(* Logix 5000 project; controller FV vendor 1 type 14 code 217 rev 31.11; software revision 31.00; part 37 of 63 *)
(* tags used below, declared in another part *)
   CWD : CHECKWORD_FLAGS;
   Dummy : BOOL;
   FV_bit_to_clear : DINT;
   FV_data_file_address : INT;
   FV_FV10C : PlantItem;   // FV10C
   FV_FV10J : PlantItem;   // FV10J
   FV_FV11C : PlantItem;   // FV11C
   FV_FV11J : PlantItem;   // FV11J
   FV_FV12C : PlantItem;   // FV12C
   FV_FV12J : PlantItem;   // FV12J
   FV_FV13C : PlantItem;   // FV13C
   FV_FV13J : PlantItem;   // FV13J
   FV_FV14C : PlantItem;   // FV14C
   FV_FV14J : PlantItem;   // FV14J
   FV_FV15C : PlantItem;   // FV15C
   FV_FV15J : PlantItem;   // FV15J
   FV_FV16C : PlantItem;   // FV16C
   FV_FV16J : PlantItem;   // FV16J
   FV_FV17C : PlantItem;   // FV17C
   FV_FV17J : PlantItem;   // FV17J
   FV_FV18C : PlantItem;   // FV18C
   FV_FV18J : PlantItem;   // FV18J
   FV_FV19C : PlantItem;   // FV19C
   FV_FV19J : PlantItem;   // FV19J
   FV_FV1C : PlantItem;   // FV1C
   FV_FV1J : PlantItem;   // FV1J
   FV_FV20C : PlantItem;   // FV20C
   FV_FV20J : PlantItem;   // FV20J
   FV_FV21C : PlantItem;   // FV21C
   FV_FV21J : PlantItem;   // FV21J
   FV_FV22C : PlantItem;   // FV22C
   FV_FV22J : PlantItem;   // FV22J
   FV_FV23C : PlantItem;   // FV23C
   FV_FV23J : PlantItem;   // FV23J
   FV_FV24C : PlantItem;   // FV24C
   FV_FV24J : PlantItem;   // FV24J
   FV_FV25C : PlantItem;   // FV25C
   FV_FV25J : PlantItem;   // FV25J
   FV_FV26C : PlantItem;   // FV26C
   FV_FV26J : PlantItem;   // FV26J
   FV_FV27C : PlantItem;   // FV27C
   FV_FV27J : PlantItem;   // FV27J
   FV_FV28C : PlantItem;   // FV28C
   FV_FV28J : PlantItem;   // FV28J
   FV_FV29C : PlantItem;   // FV29C
   FV_FV29J : PlantItem;   // FV29J
   FV_FV2C : PlantItem;   // FV2C
   FV_FV2J : PlantItem;   // FV2J
   FV_FV30C : PlantItem;   // FV30C
   FV_FV30J : PlantItem;   // FV30J
   FV_FV31C : PlantItem;   // FV31C
   FV_FV31J : PlantItem;   // FV31J
   FV_FV3C : PlantItem;   // FV3C
   FV_FV3J : PlantItem;   // FV3J
   FV_FV4C : PlantItem;   // FV4C
   FV_FV4J : PlantItem;   // FV4J
   FV_FV5C : PlantItem;   // FV5C
   FV_FV5J : PlantItem;   // FV5J
   FV_FV6C : PlantItem;   // FV6C
   FV_FV6J : PlantItem;   // FV6J
   FV_FV7C : PlantItem;   // FV7C
   FV_FV7J : PlantItem;   // FV7J
   FV_FV8C : PlantItem;   // FV8C
   FV_FV8J : PlantItem;   // FV8J
   FV_FV9C : PlantItem;   // FV9C
   FV_FV9J : PlantItem;   // FV9J
   FV_N110 : INT[255];   // FV DATA 0 CURRENT FV DATA
   FV_N111 : INT[50];   // FV1, CURRENT FV DATA
   FV_N112 : INT[50];   // FV2, CURRENT FV DATA
   FV_N113 : INT[50];   // FV3, CURRENT FV DATA
   FV_N114 : INT[50];   // FV4, CURRENT FV DATA
   FV_N115 : INT[50];   // FV5, CURRENT FV DATA
   FV_N116 : INT[50];   // FV6, CURRENT FV DATA
   FV_N117 : INT[50];   // FV7, CURRENT FV DATA
   FV_N118 : INT[50];   // FV8, CURRENT FV DATA
   FV_N119 : INT[50];   // FV9, CURRENT FV DATA
   FV_N120 : INT[50];   // FV10, CURRENT FV DATA
   FV_N121 : INT[50];   // FV11, CURRENT FV DATA
   FV_N122 : INT[50];   // FV12, CURRENT FV DATA
   FV_N123 : INT[50];   // FV13, CURRENT FV DATA
   FV_N124 : INT[50];   // FV14, CURRENT FV DATA
   FV_N125 : INT[50];   // FV15, CURRENT FV DATA
   FV_N126 : INT[50];   // FV16, CURRENT FV DATA
   FV_N127 : INT[50];   // FV17, CURRENT FV DATA
   FV_N128 : INT[50];   // FV18, CURRENT FV DATA
   FV_N129 : INT[50];   // FV19, CURRENT FV DATA
   FV_N13 : INT[255];   // PLC>ME Inter PLC comms traf fic inbound
   FV_N130 : INT[50];   // FV20, CURRENT FV DATA
   FV_N131 : INT[50];   // FV21, CURRENT FV DATA
   FV_N132 : INT[50];   // FV22, CURRENT FV DATA
   FV_N133 : INT[50];   // FV23, CURRENT FV DATA
   FV_N134 : INT[50];   // FV24, CURRENT FV DATA
   FV_N135 : INT[50];   // FV25, CURRENT FV DATA
   FV_N136 : INT[50];   // YSV1, CURRENT FV DATA
   FV_N137 : INT[50];   // YSV2, CURRENT FV DATA
   FV_N138 : INT[50];   // YSV3, CURRENT FV DATA
   FV_N139 : INT[255];   // YST1
   FV_N140 : INT[255];   // YST2
   FV_N141 : INT[255];   // YSV1 DATA
   FV_N142 : INT[255];   // YSV2 DATA
   FV_N143 : INT[255];   // YSV3 DATA
   FV_N144 : INT[255];   // YST1 DATA
   FV_N145 : INT[255];   // YST2 DATA
   FV_N146 : INT[50];   // FV26, CURRENT FV DATA
   FV_N147 : INT[50];   // FV27, CURRENT FV DATA
   FV_N148 : INT[50];   // FV28, CURRENT FV DATA
   FV_N149 : INT[50];   // FV29, CURRENT FV DATA
   FV_N150 : INT[50];   // FV30, CURRENT FV DATA
   FV_N151 : INT[50];   // FV31, CURRENT FV DATA
   FV_N210 : INT[255];   // GLYCL_PTRS
   FV_word_offset : INT;
   FV_YSV1CV : PlantItem;   // YSV1CV
   FV_YSV1J : PlantItem;   // YSV1J
   FV_YSV2CV : PlantItem;   // YSV2CV
   FV_YSV2J : PlantItem;   // YSV2J
   FV_YSV3J : PlantItem;   // YSV3J
(* FV_Common, continued *)

ROUTINE FV_Clear_Flag_In_FV_Datafile   (* ladder *)
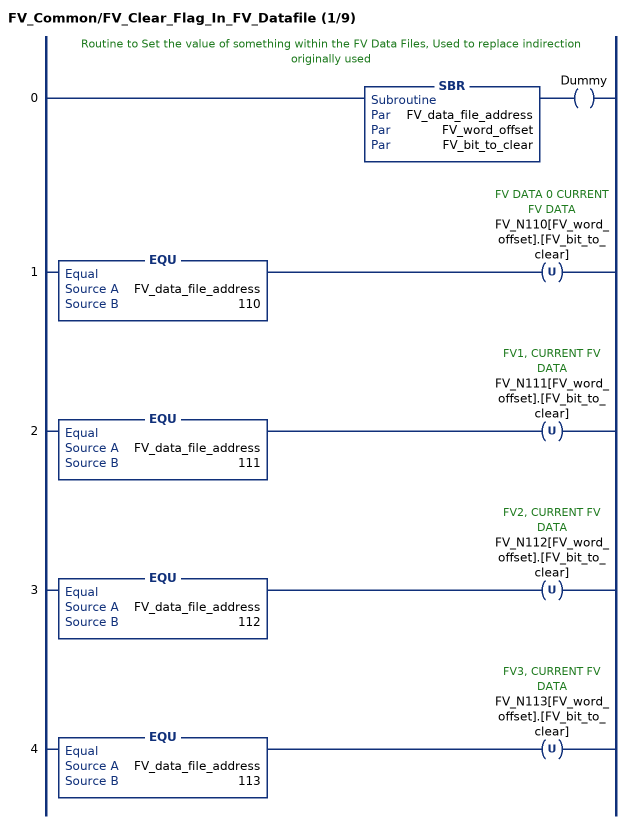
   // Routine to Set the value of something within the FV Data Files, Used to replace indirection originally used
   0: SBR(FV_data_file_address,FV_word_offset,FV_bit_to_clear)OTE(Dummy);
   1: EQU(FV_data_file_address,110)OTU(FV_N110[FV_word_offset].[FV_bit_to_clear]);
   2: EQU(FV_data_file_address,111)OTU(FV_N111[FV_word_offset].[FV_bit_to_clear]);
   3: EQU(FV_data_file_address,112)OTU(FV_N112[FV_word_offset].[FV_bit_to_clear]);
   4: EQU(FV_data_file_address,113)OTU(FV_N113[FV_word_offset].[FV_bit_to_clear]);
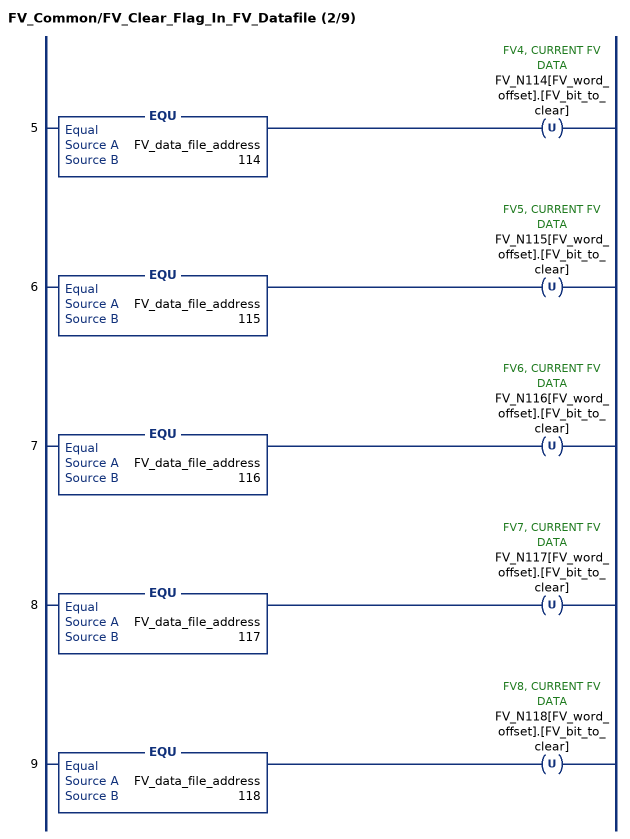
   5: EQU(FV_data_file_address,114)OTU(FV_N114[FV_word_offset].[FV_bit_to_clear]);
   6: EQU(FV_data_file_address,115)OTU(FV_N115[FV_word_offset].[FV_bit_to_clear]);
   7: EQU(FV_data_file_address,116)OTU(FV_N116[FV_word_offset].[FV_bit_to_clear]);
   8: EQU(FV_data_file_address,117)OTU(FV_N117[FV_word_offset].[FV_bit_to_clear]);
   9: EQU(FV_data_file_address,118)OTU(FV_N118[FV_word_offset].[FV_bit_to_clear]);
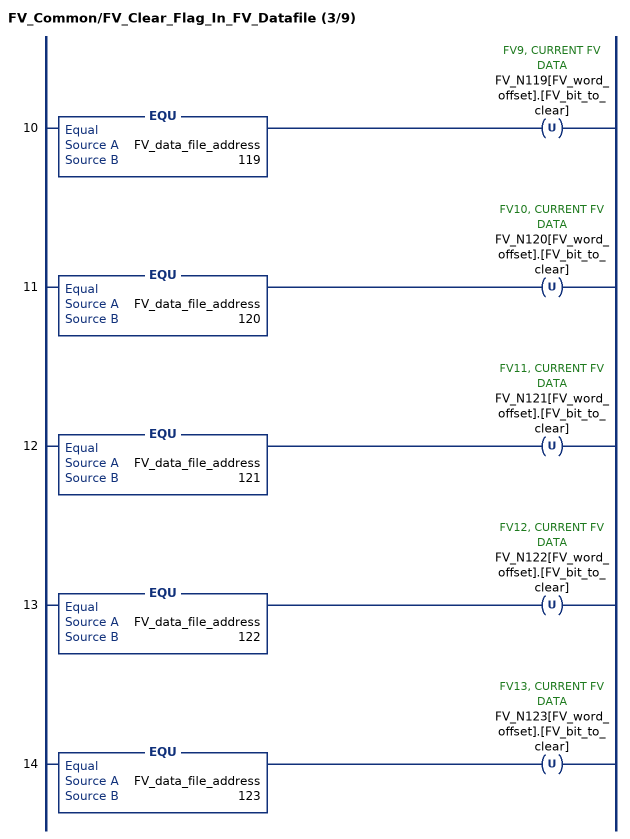
   10: EQU(FV_data_file_address,119)OTU(FV_N119[FV_word_offset].[FV_bit_to_clear]);
   11: EQU(FV_data_file_address,120)OTU(FV_N120[FV_word_offset].[FV_bit_to_clear]);
   12: EQU(FV_data_file_address,121)OTU(FV_N121[FV_word_offset].[FV_bit_to_clear]);
   13: EQU(FV_data_file_address,122)OTU(FV_N122[FV_word_offset].[FV_bit_to_clear]);
   14: EQU(FV_data_file_address,123)OTU(FV_N123[FV_word_offset].[FV_bit_to_clear]);
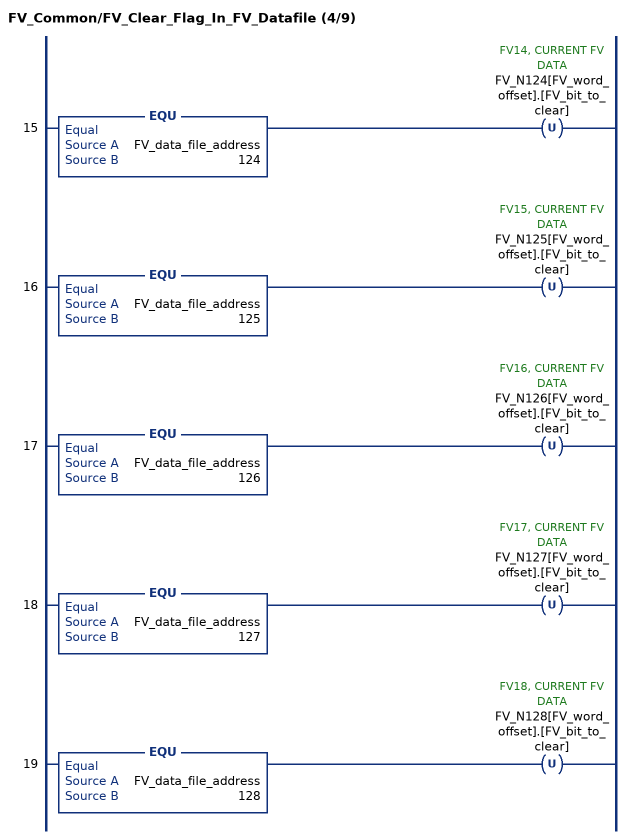
   15: EQU(FV_data_file_address,124)OTU(FV_N124[FV_word_offset].[FV_bit_to_clear]);
   16: EQU(FV_data_file_address,125)OTU(FV_N125[FV_word_offset].[FV_bit_to_clear]);
   17: EQU(FV_data_file_address,126)OTU(FV_N126[FV_word_offset].[FV_bit_to_clear]);
   18: EQU(FV_data_file_address,127)OTU(FV_N127[FV_word_offset].[FV_bit_to_clear]);
   19: EQU(FV_data_file_address,128)OTU(FV_N128[FV_word_offset].[FV_bit_to_clear]);
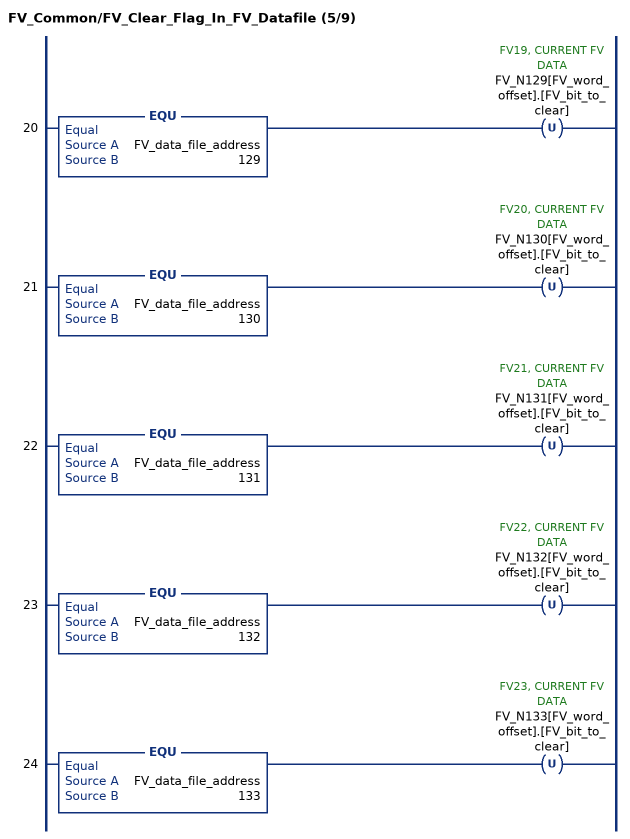
   20: EQU(FV_data_file_address,129)OTU(FV_N129[FV_word_offset].[FV_bit_to_clear]);
   21: EQU(FV_data_file_address,130)OTU(FV_N130[FV_word_offset].[FV_bit_to_clear]);
   22: EQU(FV_data_file_address,131)OTU(FV_N131[FV_word_offset].[FV_bit_to_clear]);
   23: EQU(FV_data_file_address,132)OTU(FV_N132[FV_word_offset].[FV_bit_to_clear]);
   24: EQU(FV_data_file_address,133)OTU(FV_N133[FV_word_offset].[FV_bit_to_clear]);
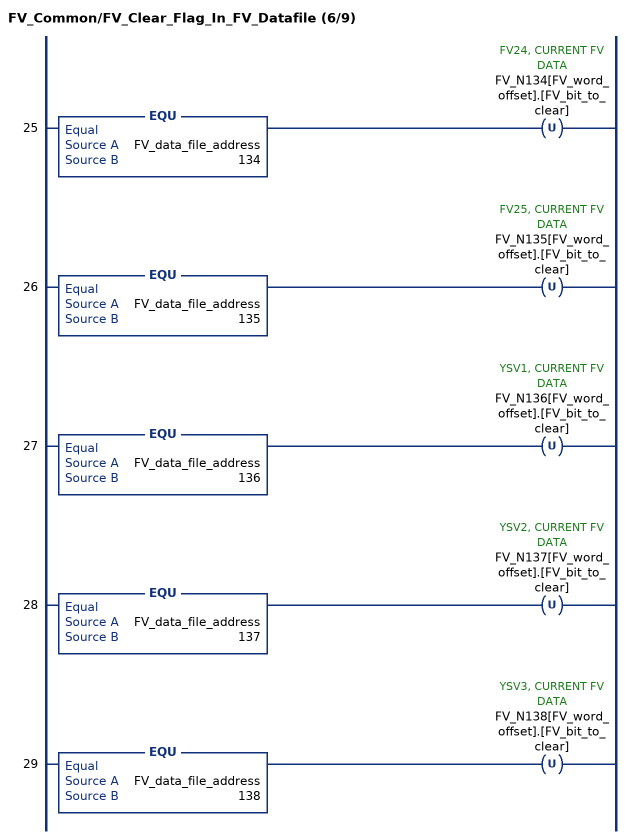
   25: EQU(FV_data_file_address,134)OTU(FV_N134[FV_word_offset].[FV_bit_to_clear]);
   26: EQU(FV_data_file_address,135)OTU(FV_N135[FV_word_offset].[FV_bit_to_clear]);
   27: EQU(FV_data_file_address,136)OTU(FV_N136[FV_word_offset].[FV_bit_to_clear]);
   28: EQU(FV_data_file_address,137)OTU(FV_N137[FV_word_offset].[FV_bit_to_clear]);
   29: EQU(FV_data_file_address,138)OTU(FV_N138[FV_word_offset].[FV_bit_to_clear]);
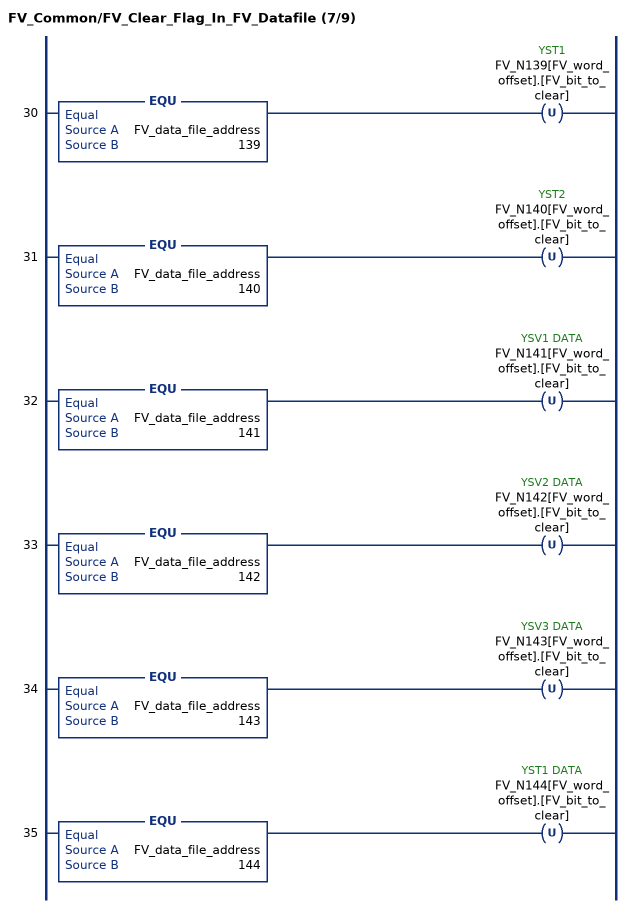
   30: EQU(FV_data_file_address,139)OTU(FV_N139[FV_word_offset].[FV_bit_to_clear]);
   31: EQU(FV_data_file_address,140)OTU(FV_N140[FV_word_offset].[FV_bit_to_clear]);
   32: EQU(FV_data_file_address,141)OTU(FV_N141[FV_word_offset].[FV_bit_to_clear]);
   33: EQU(FV_data_file_address,142)OTU(FV_N142[FV_word_offset].[FV_bit_to_clear]);
   34: EQU(FV_data_file_address,143)OTU(FV_N143[FV_word_offset].[FV_bit_to_clear]);
   35: EQU(FV_data_file_address,144)OTU(FV_N144[FV_word_offset].[FV_bit_to_clear]);
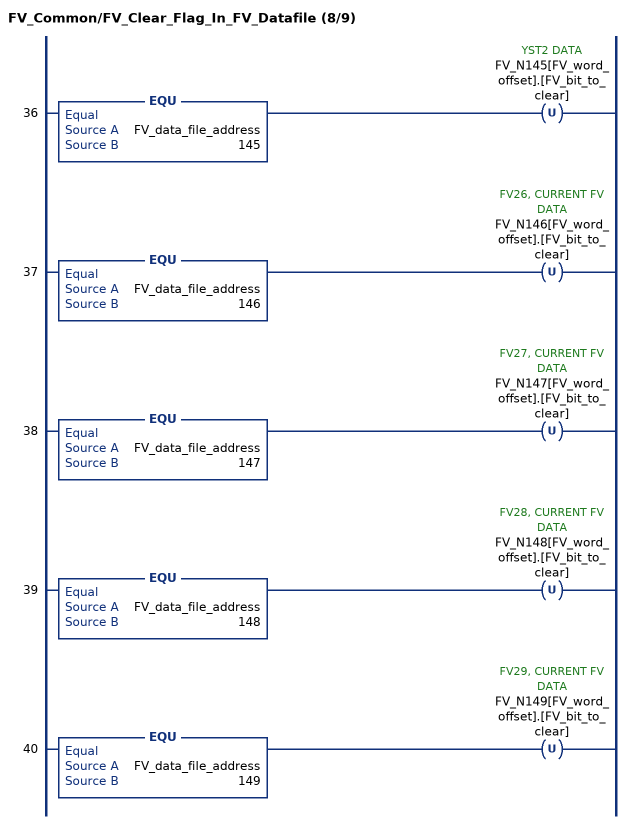
   36: EQU(FV_data_file_address,145)OTU(FV_N145[FV_word_offset].[FV_bit_to_clear]);
   37: EQU(FV_data_file_address,146)OTU(FV_N146[FV_word_offset].[FV_bit_to_clear]);
   38: EQU(FV_data_file_address,147)OTU(FV_N147[FV_word_offset].[FV_bit_to_clear]);
   39: EQU(FV_data_file_address,148)OTU(FV_N148[FV_word_offset].[FV_bit_to_clear]);
   40: EQU(FV_data_file_address,149)OTU(FV_N149[FV_word_offset].[FV_bit_to_clear]);
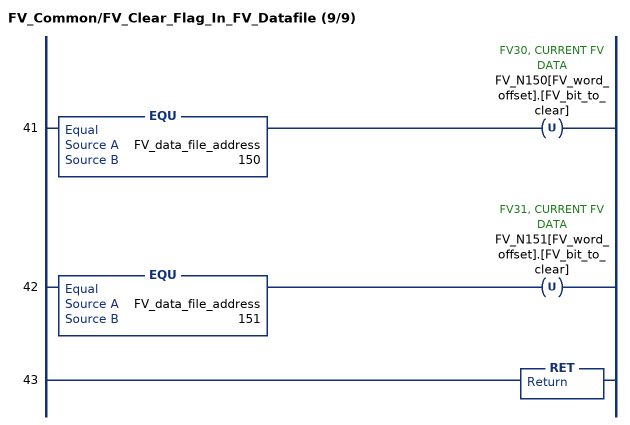
   41: EQU(FV_data_file_address,150)OTU(FV_N150[FV_word_offset].[FV_bit_to_clear]);
   42: EQU(FV_data_file_address,151)OTU(FV_N151[FV_word_offset].[FV_bit_to_clear]);
   43: RET();
END_ROUTINE

ROUTINE FV_COOLVLVOPN_111   (* ladder *)
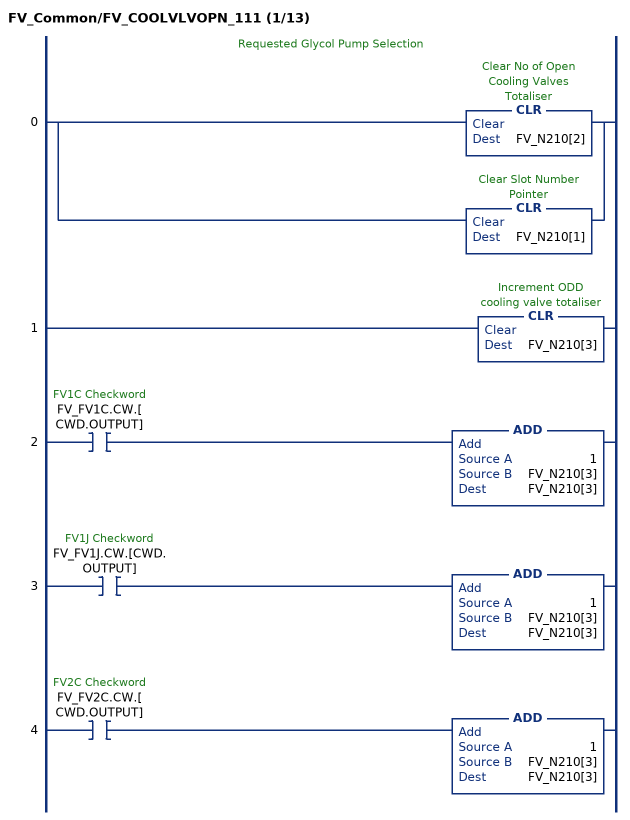
   // Requested Glycol Pump Selection
   0: [CLR(FV_N210[2]) ,CLR(FV_N210[1]) ];
   1: CLR(FV_N210[3]);
   2: XIC(FV_FV1C.CW.[CWD.OUTPUT])ADD(1,FV_N210[3],FV_N210[3]);
   3: XIC(FV_FV1J.CW.[CWD.OUTPUT])ADD(1,FV_N210[3],FV_N210[3]);
   4: XIC(FV_FV2C.CW.[CWD.OUTPUT])ADD(1,FV_N210[3],FV_N210[3]);
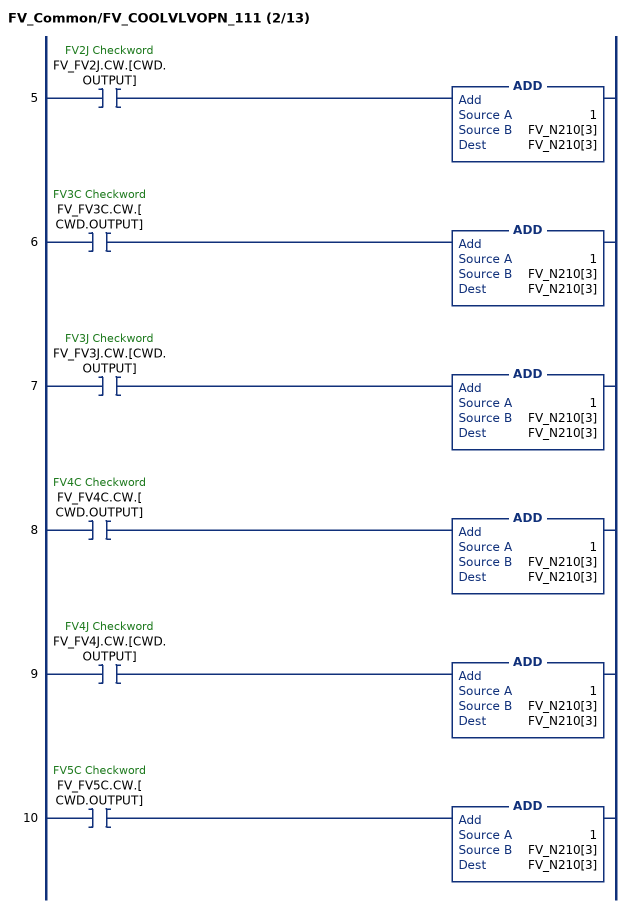
   5: XIC(FV_FV2J.CW.[CWD.OUTPUT])ADD(1,FV_N210[3],FV_N210[3]);
   6: XIC(FV_FV3C.CW.[CWD.OUTPUT])ADD(1,FV_N210[3],FV_N210[3]);
   7: XIC(FV_FV3J.CW.[CWD.OUTPUT])ADD(1,FV_N210[3],FV_N210[3]);
   8: XIC(FV_FV4C.CW.[CWD.OUTPUT])ADD(1,FV_N210[3],FV_N210[3]);
   9: XIC(FV_FV4J.CW.[CWD.OUTPUT])ADD(1,FV_N210[3],FV_N210[3]);
   10: XIC(FV_FV5C.CW.[CWD.OUTPUT])ADD(1,FV_N210[3],FV_N210[3]);
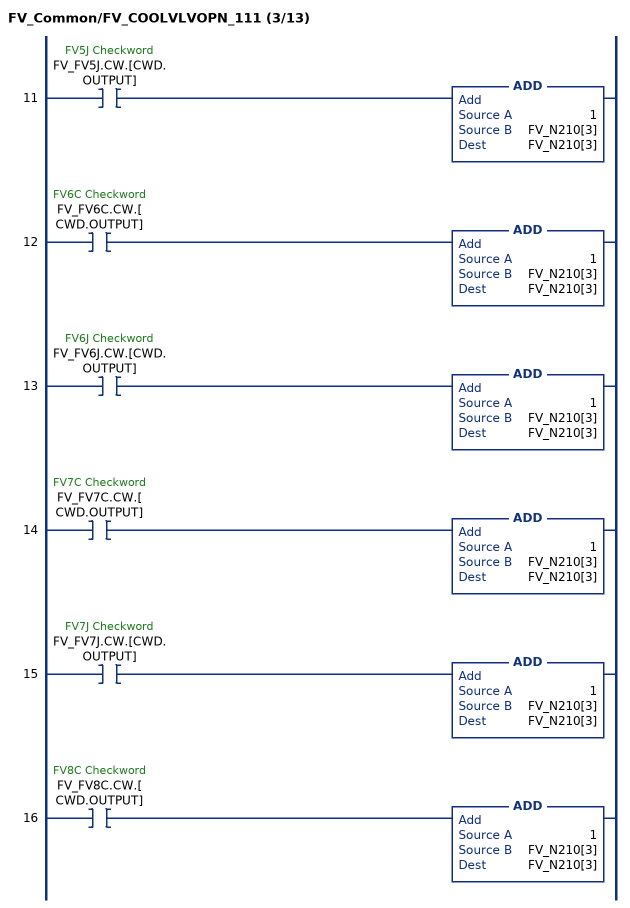
   11: XIC(FV_FV5J.CW.[CWD.OUTPUT])ADD(1,FV_N210[3],FV_N210[3]);
   12: XIC(FV_FV6C.CW.[CWD.OUTPUT])ADD(1,FV_N210[3],FV_N210[3]);
   13: XIC(FV_FV6J.CW.[CWD.OUTPUT])ADD(1,FV_N210[3],FV_N210[3]);
   14: XIC(FV_FV7C.CW.[CWD.OUTPUT])ADD(1,FV_N210[3],FV_N210[3]);
   15: XIC(FV_FV7J.CW.[CWD.OUTPUT])ADD(1,FV_N210[3],FV_N210[3]);
   16: XIC(FV_FV8C.CW.[CWD.OUTPUT])ADD(1,FV_N210[3],FV_N210[3]);
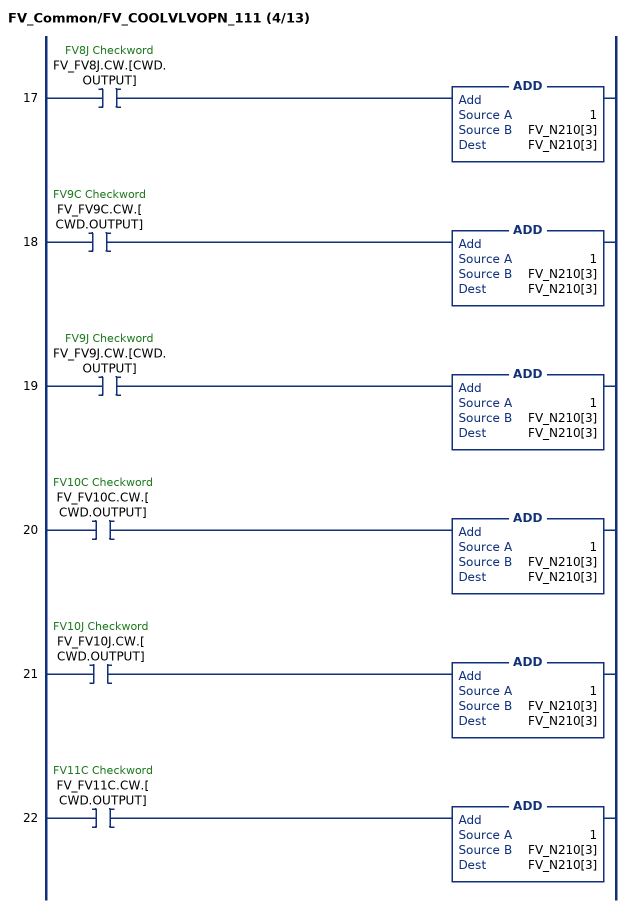
   17: XIC(FV_FV8J.CW.[CWD.OUTPUT])ADD(1,FV_N210[3],FV_N210[3]);
   18: XIC(FV_FV9C.CW.[CWD.OUTPUT])ADD(1,FV_N210[3],FV_N210[3]);
   19: XIC(FV_FV9J.CW.[CWD.OUTPUT])ADD(1,FV_N210[3],FV_N210[3]);
   20: XIC(FV_FV10C.CW.[CWD.OUTPUT])ADD(1,FV_N210[3],FV_N210[3]);
   21: XIC(FV_FV10J.CW.[CWD.OUTPUT])ADD(1,FV_N210[3],FV_N210[3]);
   22: XIC(FV_FV11C.CW.[CWD.OUTPUT])ADD(1,FV_N210[3],FV_N210[3]);
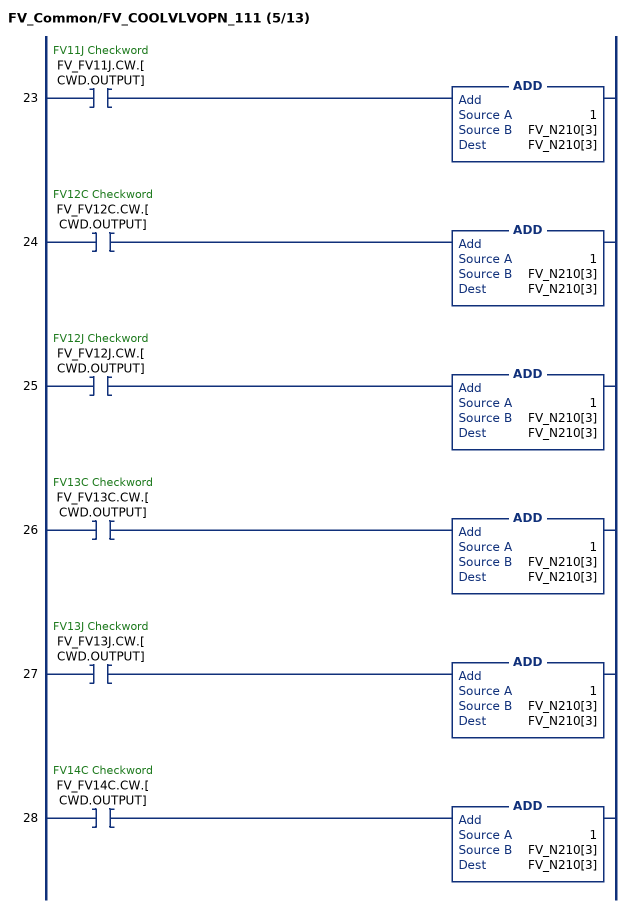
   23: XIC(FV_FV11J.CW.[CWD.OUTPUT])ADD(1,FV_N210[3],FV_N210[3]);
   24: XIC(FV_FV12C.CW.[CWD.OUTPUT])ADD(1,FV_N210[3],FV_N210[3]);
   25: XIC(FV_FV12J.CW.[CWD.OUTPUT])ADD(1,FV_N210[3],FV_N210[3]);
   26: XIC(FV_FV13C.CW.[CWD.OUTPUT])ADD(1,FV_N210[3],FV_N210[3]);
   27: XIC(FV_FV13J.CW.[CWD.OUTPUT])ADD(1,FV_N210[3],FV_N210[3]);
   28: XIC(FV_FV14C.CW.[CWD.OUTPUT])ADD(1,FV_N210[3],FV_N210[3]);
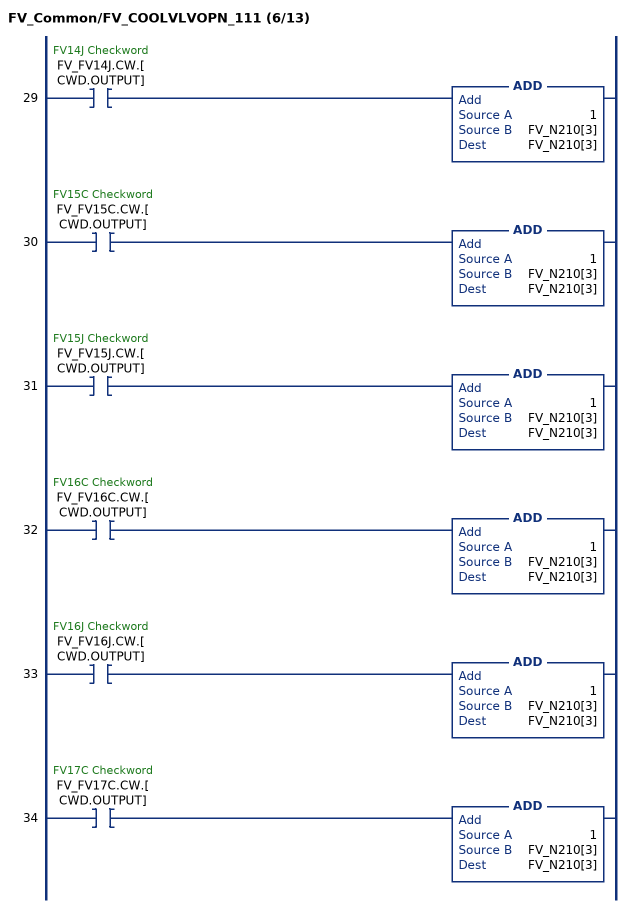
   29: XIC(FV_FV14J.CW.[CWD.OUTPUT])ADD(1,FV_N210[3],FV_N210[3]);
   30: XIC(FV_FV15C.CW.[CWD.OUTPUT])ADD(1,FV_N210[3],FV_N210[3]);
   31: XIC(FV_FV15J.CW.[CWD.OUTPUT])ADD(1,FV_N210[3],FV_N210[3]);
   32: XIC(FV_FV16C.CW.[CWD.OUTPUT])ADD(1,FV_N210[3],FV_N210[3]);
   33: XIC(FV_FV16J.CW.[CWD.OUTPUT])ADD(1,FV_N210[3],FV_N210[3]);
   34: XIC(FV_FV17C.CW.[CWD.OUTPUT])ADD(1,FV_N210[3],FV_N210[3]);
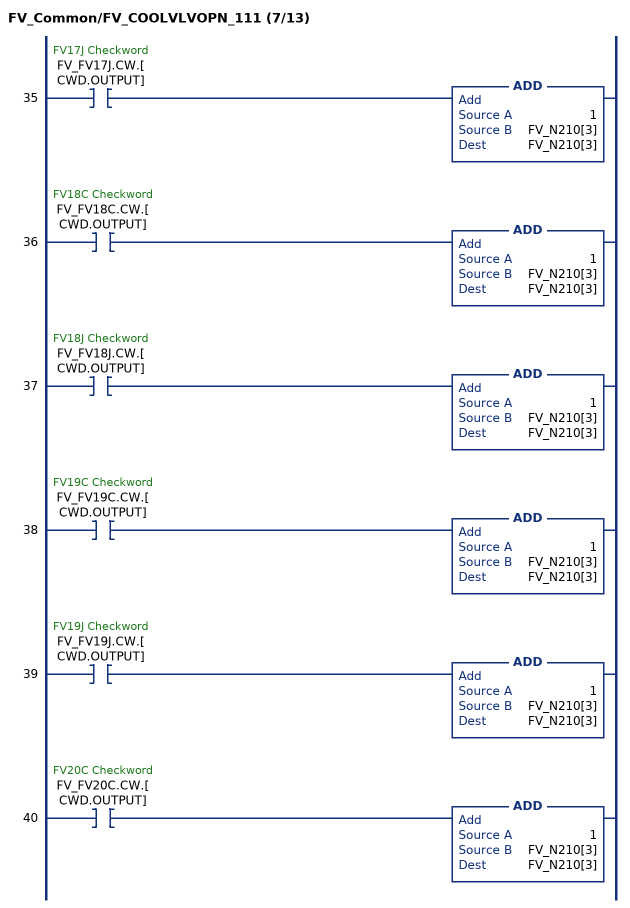
   35: XIC(FV_FV17J.CW.[CWD.OUTPUT])ADD(1,FV_N210[3],FV_N210[3]);
   36: XIC(FV_FV18C.CW.[CWD.OUTPUT])ADD(1,FV_N210[3],FV_N210[3]);
   37: XIC(FV_FV18J.CW.[CWD.OUTPUT])ADD(1,FV_N210[3],FV_N210[3]);
   38: XIC(FV_FV19C.CW.[CWD.OUTPUT])ADD(1,FV_N210[3],FV_N210[3]);
   39: XIC(FV_FV19J.CW.[CWD.OUTPUT])ADD(1,FV_N210[3],FV_N210[3]);
   40: XIC(FV_FV20C.CW.[CWD.OUTPUT])ADD(1,FV_N210[3],FV_N210[3]);
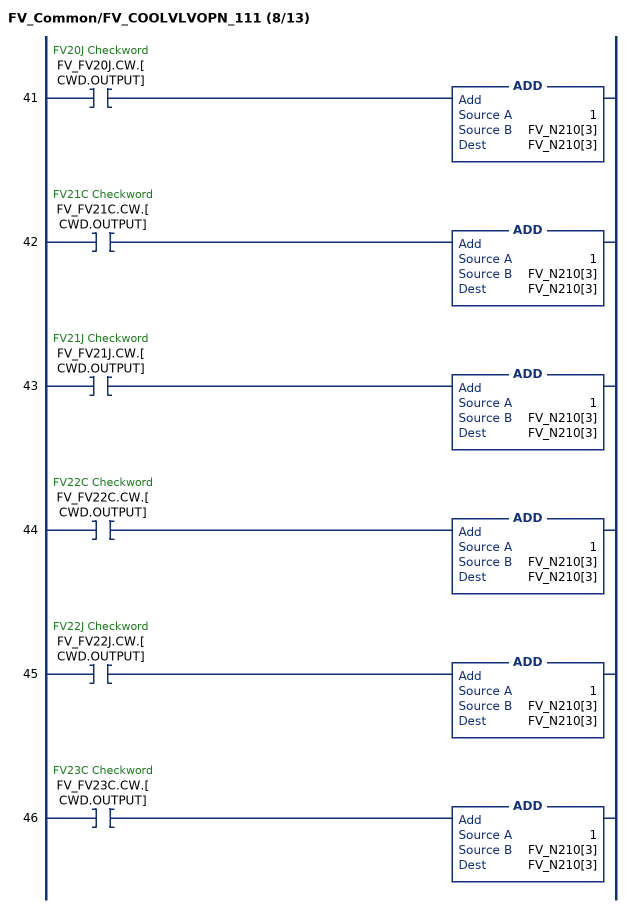
   41: XIC(FV_FV20J.CW.[CWD.OUTPUT])ADD(1,FV_N210[3],FV_N210[3]);
   42: XIC(FV_FV21C.CW.[CWD.OUTPUT])ADD(1,FV_N210[3],FV_N210[3]);
   43: XIC(FV_FV21J.CW.[CWD.OUTPUT])ADD(1,FV_N210[3],FV_N210[3]);
   44: XIC(FV_FV22C.CW.[CWD.OUTPUT])ADD(1,FV_N210[3],FV_N210[3]);
   45: XIC(FV_FV22J.CW.[CWD.OUTPUT])ADD(1,FV_N210[3],FV_N210[3]);
   46: XIC(FV_FV23C.CW.[CWD.OUTPUT])ADD(1,FV_N210[3],FV_N210[3]);
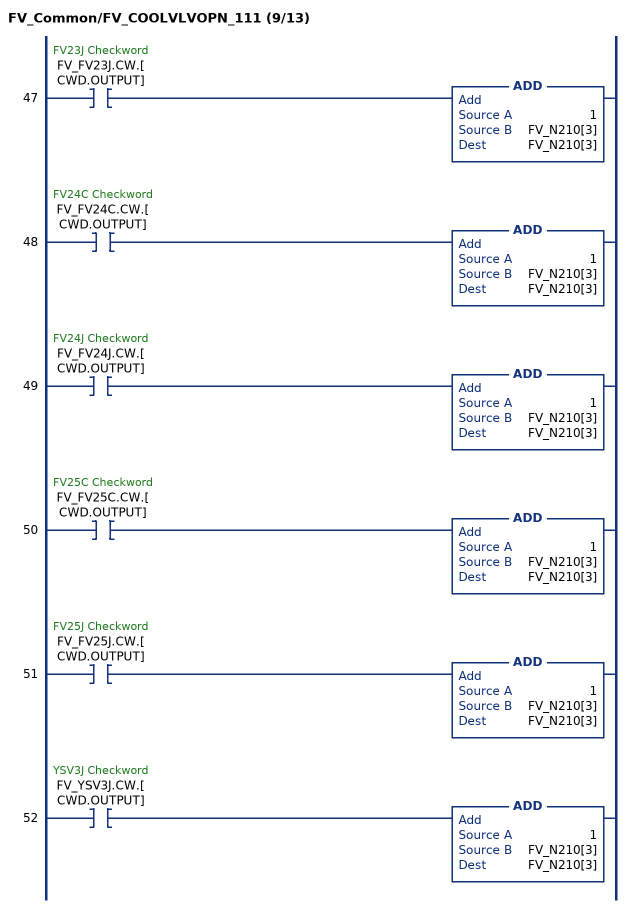
   47: XIC(FV_FV23J.CW.[CWD.OUTPUT])ADD(1,FV_N210[3],FV_N210[3]);
   48: XIC(FV_FV24C.CW.[CWD.OUTPUT])ADD(1,FV_N210[3],FV_N210[3]);
   49: XIC(FV_FV24J.CW.[CWD.OUTPUT])ADD(1,FV_N210[3],FV_N210[3]);
   50: XIC(FV_FV25C.CW.[CWD.OUTPUT])ADD(1,FV_N210[3],FV_N210[3]);
   51: XIC(FV_FV25J.CW.[CWD.OUTPUT])ADD(1,FV_N210[3],FV_N210[3]);
   52: XIC(FV_YSV3J.CW.[CWD.OUTPUT])ADD(1,FV_N210[3],FV_N210[3]);
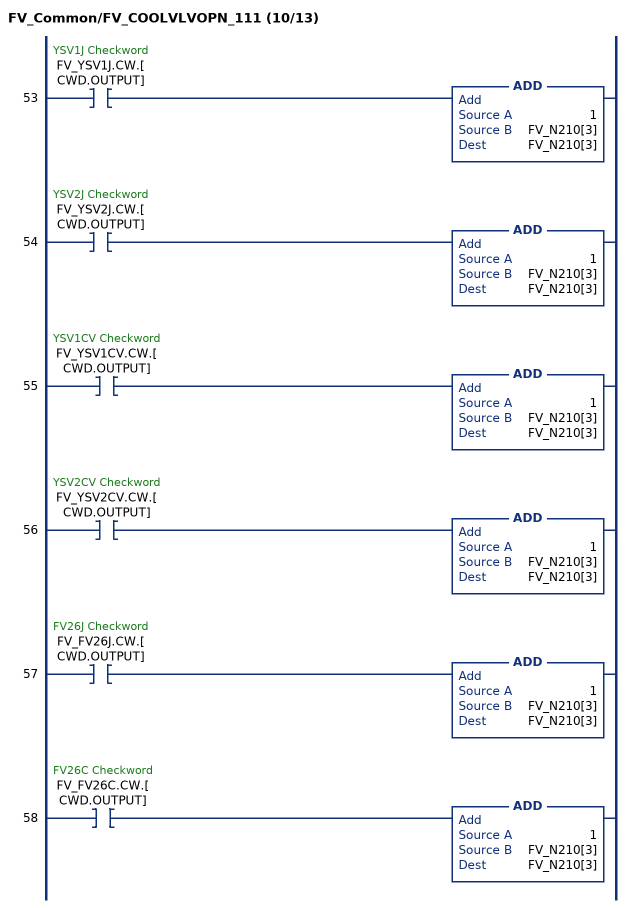
   53: XIC(FV_YSV1J.CW.[CWD.OUTPUT])ADD(1,FV_N210[3],FV_N210[3]);
   54: XIC(FV_YSV2J.CW.[CWD.OUTPUT])ADD(1,FV_N210[3],FV_N210[3]);
   55: XIC(FV_YSV1CV.CW.[CWD.OUTPUT])ADD(1,FV_N210[3],FV_N210[3]);
   56: XIC(FV_YSV2CV.CW.[CWD.OUTPUT])ADD(1,FV_N210[3],FV_N210[3]);
   57: XIC(FV_FV26J.CW.[CWD.OUTPUT])ADD(1,FV_N210[3],FV_N210[3]);
   58: XIC(FV_FV26C.CW.[CWD.OUTPUT])ADD(1,FV_N210[3],FV_N210[3]);
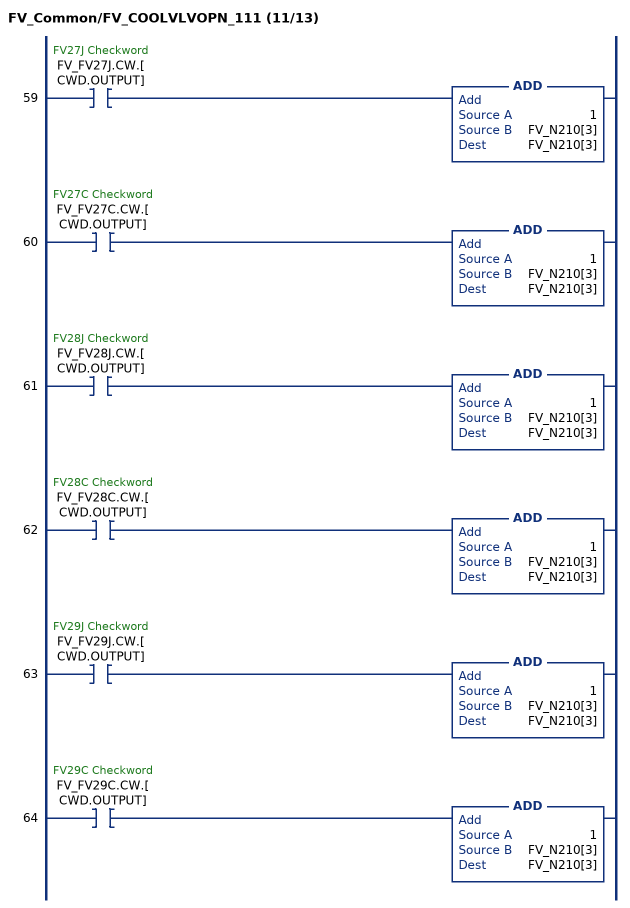
   59: XIC(FV_FV27J.CW.[CWD.OUTPUT])ADD(1,FV_N210[3],FV_N210[3]);
   60: XIC(FV_FV27C.CW.[CWD.OUTPUT])ADD(1,FV_N210[3],FV_N210[3]);
   61: XIC(FV_FV28J.CW.[CWD.OUTPUT])ADD(1,FV_N210[3],FV_N210[3]);
   62: XIC(FV_FV28C.CW.[CWD.OUTPUT])ADD(1,FV_N210[3],FV_N210[3]);
   63: XIC(FV_FV29J.CW.[CWD.OUTPUT])ADD(1,FV_N210[3],FV_N210[3]);
   64: XIC(FV_FV29C.CW.[CWD.OUTPUT])ADD(1,FV_N210[3],FV_N210[3]);
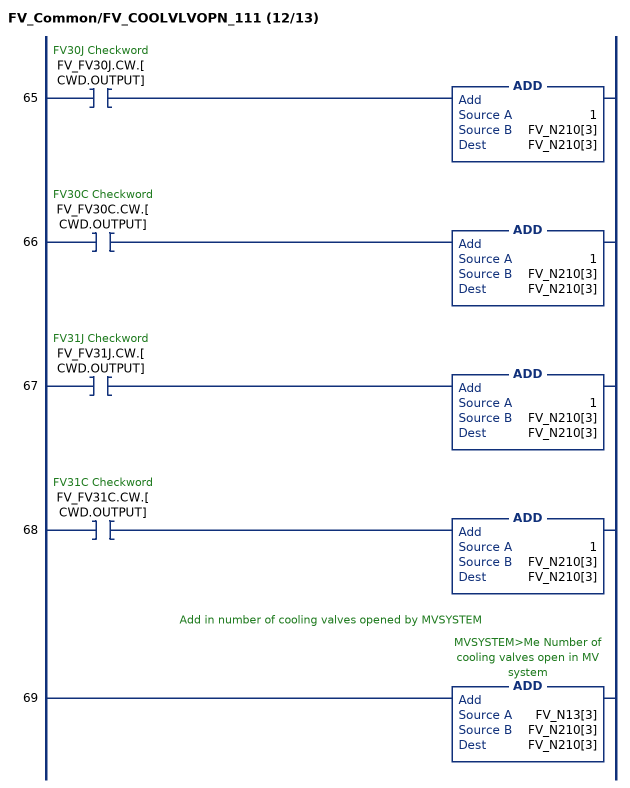
   65: XIC(FV_FV30J.CW.[CWD.OUTPUT])ADD(1,FV_N210[3],FV_N210[3]);
   66: XIC(FV_FV30C.CW.[CWD.OUTPUT])ADD(1,FV_N210[3],FV_N210[3]);
   67: XIC(FV_FV31J.CW.[CWD.OUTPUT])ADD(1,FV_N210[3],FV_N210[3]);
   68: XIC(FV_FV31C.CW.[CWD.OUTPUT])ADD(1,FV_N210[3],FV_N210[3]);
   // Add in number of cooling valves opened by MVSYSTEM
   69: ADD(FV_N13[3],FV_N210[3],FV_N210[3]);
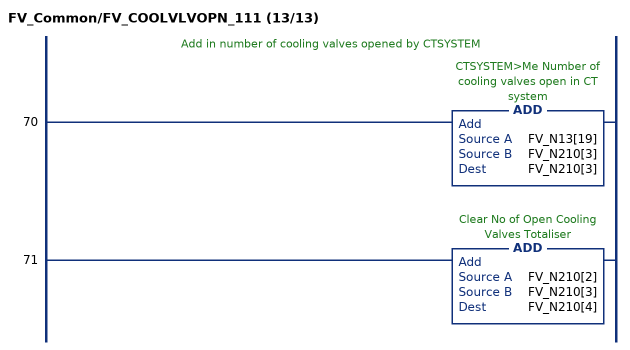
   // Add in number of cooling valves opened by CTSYSTEM
   70: ADD(FV_N13[19],FV_N210[3],FV_N210[3]);
   71: ADD(FV_N210[2],FV_N210[3],FV_N210[4]);
END_ROUTINE
